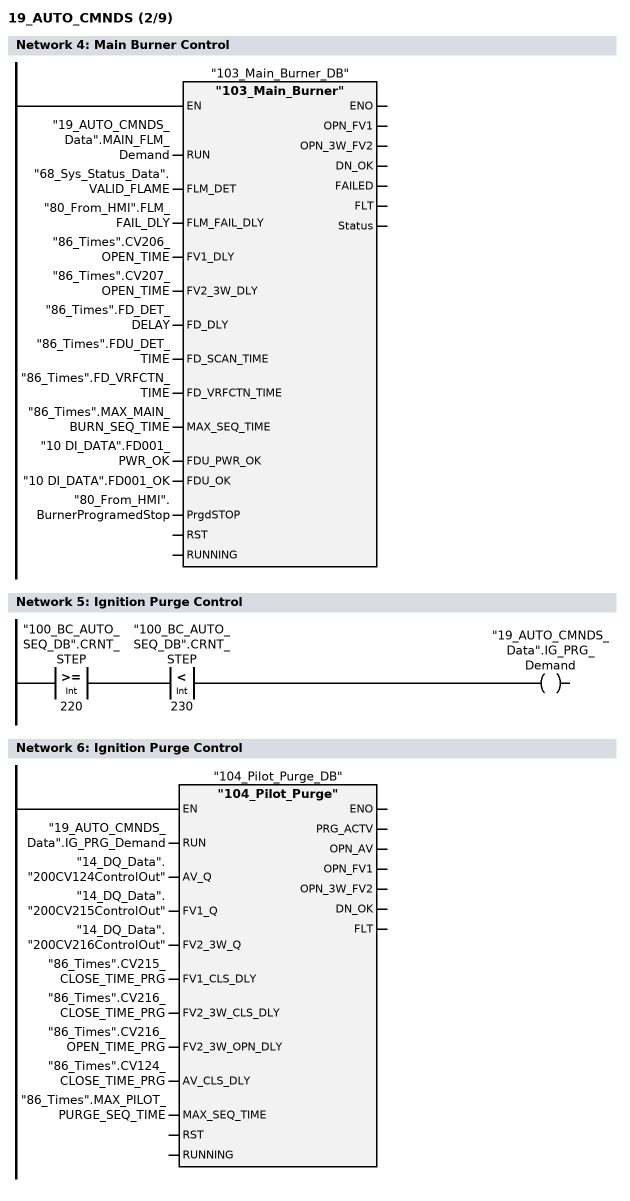
   RUNG wire#powerrail
      "103_Main_Burner_DB"(RUN := "19_AUTO_CMNDS_Data".MAIN_FLM_Demand, FLM_DET := "68_Sys_Status_Data".VALID_FLAME, FLM_FAIL_DLY := "80_From_HMI".FLM_FAIL_DLY, FV1_DLY := "86_Times".CV206_OPEN_TIME, FV2_3W_DLY := "86_Times".CV207_OPEN_TIME, FD_DLY := "86_Times".FD_DET_DELAY, FD_SCAN_TIME := "86_Times".FDU_DET_TIME, FD_VRFCTN_TIME := "86_Times".FD_VRFCTN_TIME, MAX_SEQ_TIME := "86_Times".MAX_MAIN_BURN_SEQ_TIME, FDU_PWR_OK := "10 DI_DATA".FD001_PWR_OK, FDU_OK := "10 DI_DATA".FD001_OK, PrgdSTOP := "80_From_HMI".BurnerProgramedStop, RST :=, RUNNING :=, OPN_FV1 =>, OPN_3W_FV2 =>, DN_OK =>, FAILED =>, FLT =>, Status =>)
   END_RUNG
   // the same network as SCL:
   "103_Main_Burner_DB"(RUN := "19_AUTO_CMNDS_Data".MAIN_FLM_Demand,   // "103_Main_Burner"
                        FLM_DET := "68_Sys_Status_Data".VALID_FLAME,
                        FLM_FAIL_DLY := "80_From_HMI".FLM_FAIL_DLY,
                        FV1_DLY := "86_Times".CV206_OPEN_TIME,
                        FV2_3W_DLY := "86_Times".CV207_OPEN_TIME,
                        FD_DLY := "86_Times".FD_DET_DELAY,
                        FD_SCAN_TIME := "86_Times".FDU_DET_TIME,
                        FD_VRFCTN_TIME := "86_Times".FD_VRFCTN_TIME,
                        MAX_SEQ_TIME := "86_Times".MAX_MAIN_BURN_SEQ_TIME,
                        FDU_PWR_OK := "10 DI_DATA".FD001_PWR_OK,
                        FDU_OK := "10 DI_DATA".FD001_OK,
                        PrgdSTOP := "80_From_HMI".BurnerProgramedStop);
END_REGION

REGION Network 5: Ignition Purge Control
   RUNG wire#powerrail
      { S7_Templates := "SrcType := Int" } GE_Contact(in1 := "100_BC_AUTO_SEQ_DB".CRNT_STEP, in2 := 220)
      { S7_Templates := "SrcType := Int" } LT_Contact(in1 := "100_BC_AUTO_SEQ_DB".CRNT_STEP, in2 := 230)
      Coil( "19_AUTO_CMNDS_Data".IG_PRG_Demand )
   END_RUNG
   // the same network as SCL:
   "19_AUTO_CMNDS_Data".IG_PRG_Demand := ("100_BC_AUTO_SEQ_DB".CRNT_STEP >= 220) AND ("100_BC_AUTO_SEQ_DB".CRNT_STEP < 230);
END_REGION

REGION Network 6: Ignition Purge Control
   RUNG wire#powerrail
      "104_Pilot_Purge_DB"(RUN := "19_AUTO_CMNDS_Data".IG_PRG_Demand, AV_Q := "14_DQ_Data"."200CV124ControlOut", FV1_Q := "14_DQ_Data"."200CV215ControlOut", FV2_3W_Q := "14_DQ_Data"."200CV216ControlOut", FV1_CLS_DLY := "86_Times".CV215_CLOSE_TIME_PRG, FV2_3W_CLS_DLY := "86_Times".CV216_CLOSE_TIME_PRG, FV2_3W_OPN_DLY := "86_Times".CV216_OPEN_TIME_PRG, AV_CLS_DLY := "86_Times".CV124_CLOSE_TIME_PRG, MAX_SEQ_TIME := "86_Times".MAX_PILOT_PURGE_SEQ_TIME, RST :=, RUNNING :=, PRG_ACTV =>, OPN_AV =>, OPN_FV1 =>, OPN_3W_FV2 =>, DN_OK =>, FLT =>)
   END_RUNG
   // the same network as SCL:
   "104_Pilot_Purge_DB"(RUN := "19_AUTO_CMNDS_Data".IG_PRG_Demand,   // "104_Pilot_Purge"
                        AV_Q := "14_DQ_Data"."200CV124ControlOut",
                        FV1_Q := "14_DQ_Data"."200CV215ControlOut",
                        FV2_3W_Q := "14_DQ_Data"."200CV216ControlOut",
                        FV1_CLS_DLY := "86_Times".CV215_CLOSE_TIME_PRG,
                        FV2_3W_CLS_DLY := "86_Times".CV216_CLOSE_TIME_PRG,
                        FV2_3W_OPN_DLY := "86_Times".CV216_OPEN_TIME_PRG,
                        AV_CLS_DLY := "86_Times".CV124_CLOSE_TIME_PRG,
                        MAX_SEQ_TIME := "86_Times".MAX_PILOT_PURGE_SEQ_TIME);
END_REGION

REGION Network 7: Q0.0 - Test pressure valve control CV127
   // True = Open, False = Closed
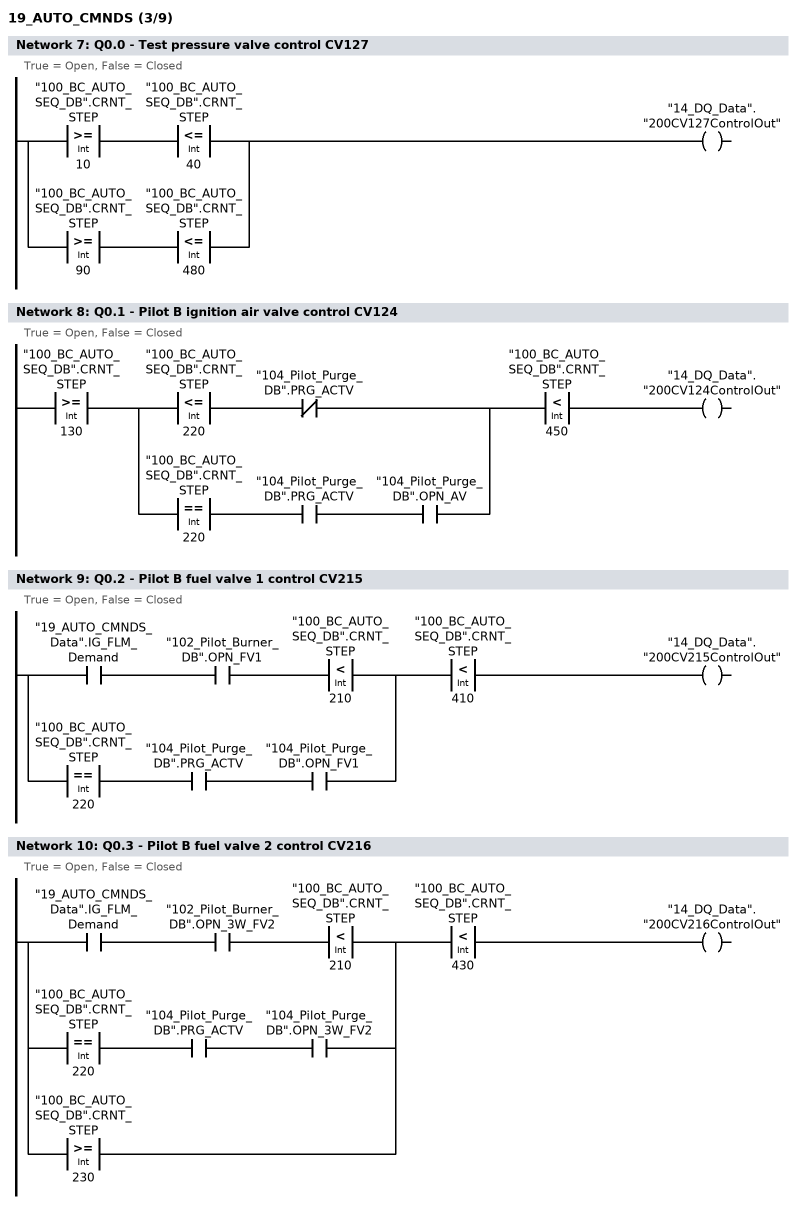
   RUNG wire#powerrail
      { S7_Templates := "SrcType := Int" } GE_Contact(in1 := "100_BC_AUTO_SEQ_DB".CRNT_STEP, in2 := 10)
      { S7_Templates := "SrcType := Int" } LE_Contact(in1 := "100_BC_AUTO_SEQ_DB".CRNT_STEP, in2 := 40)
      wire#w1
      Coil( "14_DQ_Data"."200CV127ControlOut" )
   END_RUNG
   RUNG wire#powerrail
      { S7_Templates := "SrcType := Int" } GE_Contact(in1 := "100_BC_AUTO_SEQ_DB".CRNT_STEP, in2 := 90)
      { S7_Templates := "SrcType := Int" } LE_Contact(in1 := "100_BC_AUTO_SEQ_DB".CRNT_STEP, in2 := 480)
   END_RUNG wire#w1
   // the same network as SCL:
   "14_DQ_Data"."200CV127ControlOut" := (("100_BC_AUTO_SEQ_DB".CRNT_STEP >= 10) AND ("100_BC_AUTO_SEQ_DB".CRNT_STEP <= 40)) OR (("100_BC_AUTO_SEQ_DB".CRNT_STEP >= 90) AND ("100_BC_AUTO_SEQ_DB".CRNT_STEP <= 480));
END_REGION

REGION Network 8: Q0.1 - Pilot B ignition air valve control CV124
   // True = Open, False = Closed
   RUNG wire#powerrail
      { S7_Templates := "SrcType := Int" } GE_Contact(in1 := "100_BC_AUTO_SEQ_DB".CRNT_STEP, in2 := 130)
      wire#w1
      { S7_Templates := "SrcType := Int" } LE_Contact(in1 := "100_BC_AUTO_SEQ_DB".CRNT_STEP, in2 := 220)
      I_Contact( "104_Pilot_Purge_DB".PRG_ACTV )
      wire#w2
      { S7_Templates := "SrcType := Int" } LT_Contact(in1 := "100_BC_AUTO_SEQ_DB".CRNT_STEP, in2 := 450)
      Coil( "14_DQ_Data"."200CV124ControlOut" )
   END_RUNG
   RUNG wire#w1
      { S7_Templates := "SrcType := Int" } EQ_Contact(in1 := "100_BC_AUTO_SEQ_DB".CRNT_STEP, in2 := 220)
      Contact( "104_Pilot_Purge_DB".PRG_ACTV )
      Contact( "104_Pilot_Purge_DB".OPN_AV )
   END_RUNG wire#w2
   // the same network as SCL:
   "14_DQ_Data"."200CV124ControlOut" := ("100_BC_AUTO_SEQ_DB".CRNT_STEP >= 130) AND ((("100_BC_AUTO_SEQ_DB".CRNT_STEP <= 220) AND NOT "104_Pilot_Purge_DB".PRG_ACTV) OR (("100_BC_AUTO_SEQ_DB".CRNT_STEP = 220) AND "104_Pilot_Purge_DB".PRG_ACTV AND "104_Pilot_Purge_DB".OPN_AV)) AND ("100_BC_AUTO_SEQ_DB".CRNT_STEP < 450);
END_REGION

REGION Network 9: Q0.2 - Pilot B fuel valve 1 control CV215
   // True = Open, False = Closed
   RUNG wire#powerrail
      Contact( "19_AUTO_CMNDS_Data".IG_FLM_Demand )
      Contact( "102_Pilot_Burner_DB".OPN_FV1 )
      { S7_Templates := "SrcType := Int" } LT_Contact(in1 := "100_BC_AUTO_SEQ_DB".CRNT_STEP, in2 := 210)
      wire#w1
      { S7_Templates := "SrcType := Int" } LT_Contact(in1 := "100_BC_AUTO_SEQ_DB".CRNT_STEP, in2 := 410)
      Coil( "14_DQ_Data"."200CV215ControlOut" )
   END_RUNG
   RUNG wire#powerrail
      { S7_Templates := "SrcType := Int" } EQ_Contact(in1 := "100_BC_AUTO_SEQ_DB".CRNT_STEP, in2 := 220)
      Contact( "104_Pilot_Purge_DB".PRG_ACTV )
      Contact( "104_Pilot_Purge_DB".OPN_FV1 )
   END_RUNG wire#w1
   // the same network as SCL:
   "14_DQ_Data"."200CV215ControlOut" := (("19_AUTO_CMNDS_Data".IG_FLM_Demand AND "102_Pilot_Burner_DB".OPN_FV1 AND ("100_BC_AUTO_SEQ_DB".CRNT_STEP < 210)) OR (("100_BC_AUTO_SEQ_DB".CRNT_STEP = 220) AND "104_Pilot_Purge_DB".PRG_ACTV AND "104_Pilot_Purge_DB".OPN_FV1)) AND ("100_BC_AUTO_SEQ_DB".CRNT_STEP < 410);
END_REGION

REGION Network 10: Q0.3 - Pilot B fuel valve 2 control CV216
   // True = Open, False = Closed
   RUNG wire#powerrail
      Contact( "19_AUTO_CMNDS_Data".IG_FLM_Demand )
      Contact( "102_Pilot_Burner_DB".OPN_3W_FV2 )
      { S7_Templates := "SrcType := Int" } LT_Contact(in1 := "100_BC_AUTO_SEQ_DB".CRNT_STEP, in2 := 210)
      wire#w1
      { S7_Templates := "SrcType := Int" } LT_Contact(in1 := "100_BC_AUTO_SEQ_DB".CRNT_STEP, in2 := 430)
      Coil( "14_DQ_Data"."200CV216ControlOut" )
   END_RUNG
   RUNG wire#powerrail
      { S7_Templates := "SrcType := Int" } EQ_Contact(in1 := "100_BC_AUTO_SEQ_DB".CRNT_STEP, in2 := 220)
      Contact( "104_Pilot_Purge_DB".PRG_ACTV )
      Contact( "104_Pilot_Purge_DB".OPN_3W_FV2 )
   END_RUNG wire#w1
   RUNG wire#powerrail
      { S7_Templates := "SrcType := Int" } GE_Contact(in1 := "100_BC_AUTO_SEQ_DB".CRNT_STEP, in2 := 230)
   END_RUNG wire#w1
   // the same network as SCL:
   "14_DQ_Data"."200CV216ControlOut" := (("19_AUTO_CMNDS_Data".IG_FLM_Demand AND "102_Pilot_Burner_DB".OPN_3W_FV2 AND ("100_BC_AUTO_SEQ_DB".CRNT_STEP < 210)) OR (("100_BC_AUTO_SEQ_DB".CRNT_STEP = 220) AND "104_Pilot_Purge_DB".PRG_ACTV AND "104_Pilot_Purge_DB".OPN_3W_FV2) OR ("100_BC_AUTO_SEQ_DB".CRNT_STEP >= 230)) AND ("100_BC_AUTO_SEQ_DB".CRNT_STEP < 430);
END_REGION

REGION Network 11: Q0.4 - Main B atom air valve control CV114
   // True = Open, False = Closed
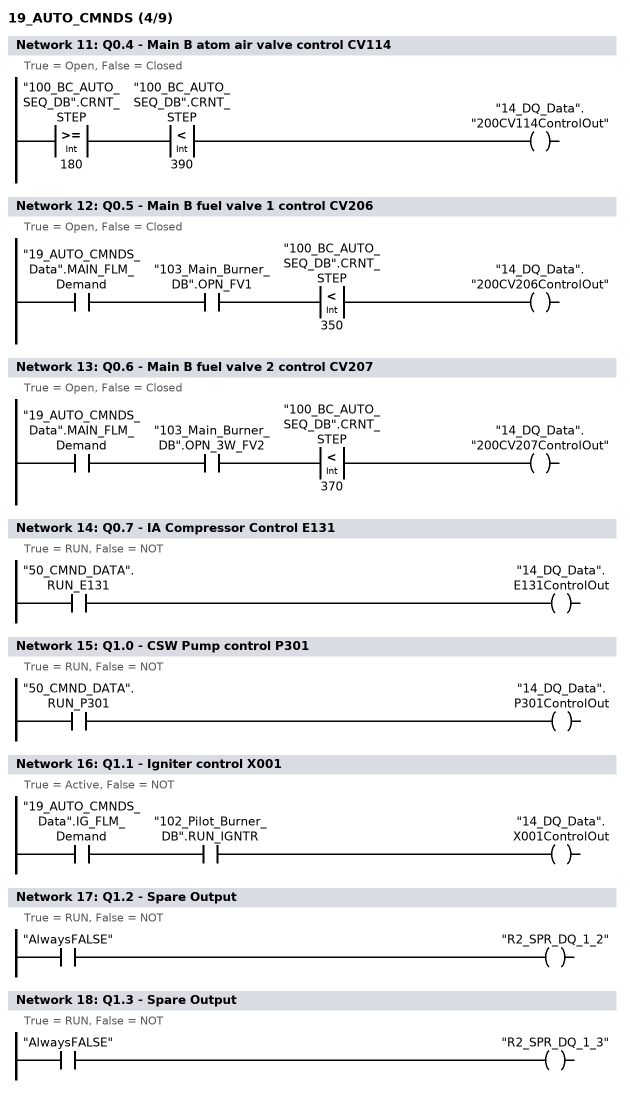
   RUNG wire#powerrail
      { S7_Templates := "SrcType := Int" } GE_Contact(in1 := "100_BC_AUTO_SEQ_DB".CRNT_STEP, in2 := 180)
      { S7_Templates := "SrcType := Int" } LT_Contact(in1 := "100_BC_AUTO_SEQ_DB".CRNT_STEP, in2 := 390)
      Coil( "14_DQ_Data"."200CV114ControlOut" )
   END_RUNG
   // the same network as SCL:
   "14_DQ_Data"."200CV114ControlOut" := ("100_BC_AUTO_SEQ_DB".CRNT_STEP >= 180) AND ("100_BC_AUTO_SEQ_DB".CRNT_STEP < 390);
END_REGION

REGION Network 12: Q0.5 - Main B fuel valve 1 control CV206
   // True = Open, False = Closed
   RUNG wire#powerrail
      Contact( "19_AUTO_CMNDS_Data".MAIN_FLM_Demand )
      Contact( "103_Main_Burner_DB".OPN_FV1 )
      { S7_Templates := "SrcType := Int" } LT_Contact(in1 := "100_BC_AUTO_SEQ_DB".CRNT_STEP, in2 := 350)
      Coil( "14_DQ_Data"."200CV206ControlOut" )
   END_RUNG
   // the same network as SCL:
   "14_DQ_Data"."200CV206ControlOut" := "19_AUTO_CMNDS_Data".MAIN_FLM_Demand AND "103_Main_Burner_DB".OPN_FV1 AND ("100_BC_AUTO_SEQ_DB".CRNT_STEP < 350);
END_REGION

REGION Network 13: Q0.6 - Main B fuel valve 2 control CV207
   // True = Open, False = Closed
   RUNG wire#powerrail
      Contact( "19_AUTO_CMNDS_Data".MAIN_FLM_Demand )
      Contact( "103_Main_Burner_DB".OPN_3W_FV2 )
      { S7_Templates := "SrcType := Int" } LT_Contact(in1 := "100_BC_AUTO_SEQ_DB".CRNT_STEP, in2 := 370)
      Coil( "14_DQ_Data"."200CV207ControlOut" )
   END_RUNG
   // the same network as SCL:
   "14_DQ_Data"."200CV207ControlOut" := "19_AUTO_CMNDS_Data".MAIN_FLM_Demand AND "103_Main_Burner_DB".OPN_3W_FV2 AND ("100_BC_AUTO_SEQ_DB".CRNT_STEP < 370);
END_REGION

REGION Network 14: Q0.7 - IA Compressor Control E131
   // True = RUN, False = NOT
   RUNG wire#powerrail
      Contact( "50_CMND_DATA".RUN_E131 )
      Coil( "14_DQ_Data".E131ControlOut )
   END_RUNG
   // the same network as SCL:
   "14_DQ_Data".E131ControlOut := "50_CMND_DATA".RUN_E131;
END_REGION

REGION Network 15: Q1.0 - CSW Pump control P301
   // True = RUN, False = NOT
   RUNG wire#powerrail
      Contact( "50_CMND_DATA".RUN_P301 )
      Coil( "14_DQ_Data".P301ControlOut )
   END_RUNG
   // the same network as SCL:
   "14_DQ_Data".P301ControlOut := "50_CMND_DATA".RUN_P301;
END_REGION

REGION Network 16: Q1.1 - Igniter control X001
   // True = Active, False = NOT
   RUNG wire#powerrail
      Contact( "19_AUTO_CMNDS_Data".IG_FLM_Demand )
      Contact( "102_Pilot_Burner_DB".RUN_IGNTR )
      Coil( "14_DQ_Data".X001ControlOut )
   END_RUNG
   // the same network as SCL:
   "14_DQ_Data".X001ControlOut := "19_AUTO_CMNDS_Data".IG_FLM_Demand AND "102_Pilot_Burner_DB".RUN_IGNTR;
END_REGION

REGION Network 17: Q1.2 - Spare Output
   // True = RUN, False = NOT
   RUNG wire#powerrail
      Contact( "AlwaysFALSE" )
      Coil( "R2_SPR_DQ_1_2" )
   END_RUNG
   // the same network as SCL:
   "R2_SPR_DQ_1_2" := "AlwaysFALSE";
END_REGION

REGION Network 18: Q1.3 - Spare Output
   // True = RUN, False = NOT
   RUNG wire#powerrail
      Contact( "AlwaysFALSE" )
      Coil( "R2_SPR_DQ_1_3" )
   END_RUNG
   // the same network as SCL:
   "R2_SPR_DQ_1_3" := "AlwaysFALSE";
END_REGION

REGION Network 19: Q1.4 - Spare Output
   // True = RUN, False = NOT
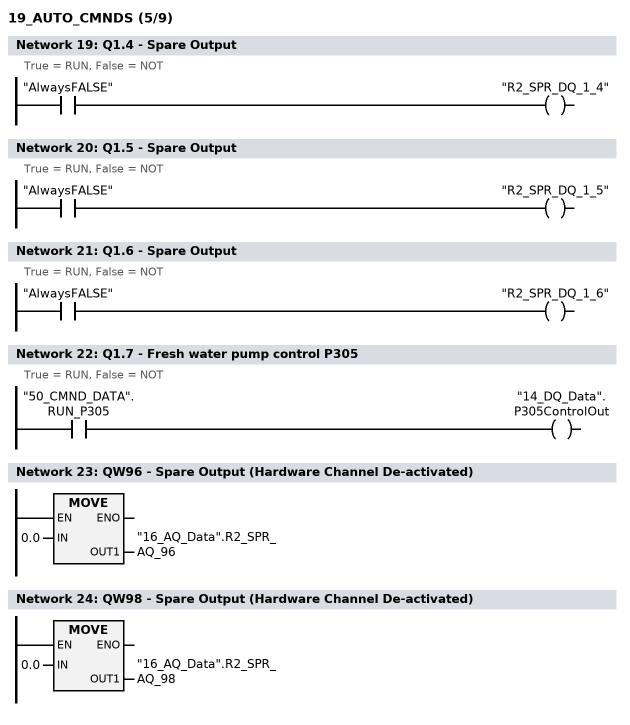
   RUNG wire#powerrail
      Contact( "AlwaysFALSE" )
      Coil( "R2_SPR_DQ_1_4" )
   END_RUNG
   // the same network as SCL:
   "R2_SPR_DQ_1_4" := "AlwaysFALSE";
END_REGION

REGION Network 20: Q1.5 - Spare Output
   // True = RUN, False = NOT
   RUNG wire#powerrail
      Contact( "AlwaysFALSE" )
      Coil( "R2_SPR_DQ_1_5" )
   END_RUNG
   // the same network as SCL:
   "R2_SPR_DQ_1_5" := "AlwaysFALSE";
END_REGION

REGION Network 21: Q1.6 - Spare Output
   // True = RUN, False = NOT
   RUNG wire#powerrail
      Contact( "AlwaysFALSE" )
      Coil( "R2_SPR_DQ_1_6" )
   END_RUNG
   // the same network as SCL:
   "R2_SPR_DQ_1_6" := "AlwaysFALSE";
END_REGION

REGION Network 22: Q1.7 - Fresh water pump control P305
   // True = RUN, False = NOT
   RUNG wire#powerrail
      Contact( "50_CMND_DATA".RUN_P305 )
      Coil( "14_DQ_Data".P305ControlOut )
   END_RUNG
   // the same network as SCL:
   "14_DQ_Data".P305ControlOut := "50_CMND_DATA".RUN_P305;
END_REGION

REGION Network 23: QW96 - Spare Output (Hardware Channel De-activated)
   RUNG wire#powerrail
      Move(in := 0.0, out1 => "16_AQ_Data".R2_SPR_AQ_96)
   END_RUNG
   // the same network as SCL:
   "16_AQ_Data".R2_SPR_AQ_96 := 0.0;
END_REGION

REGION Network 24: QW98 - Spare Output (Hardware Channel De-activated)
   RUNG wire#powerrail
      Move(in := 0.0, out1 => "16_AQ_Data".R2_SPR_AQ_98)
   END_RUNG
   // the same network as SCL:
   "16_AQ_Data".R2_SPR_AQ_98 := 0.0;
END_REGION

REGION Network 25: QW100 - Main Fuel Reg Valve Control CV203 (For Main Burn Start)
   // Changed from 20 to 230 at 160 to230 for test
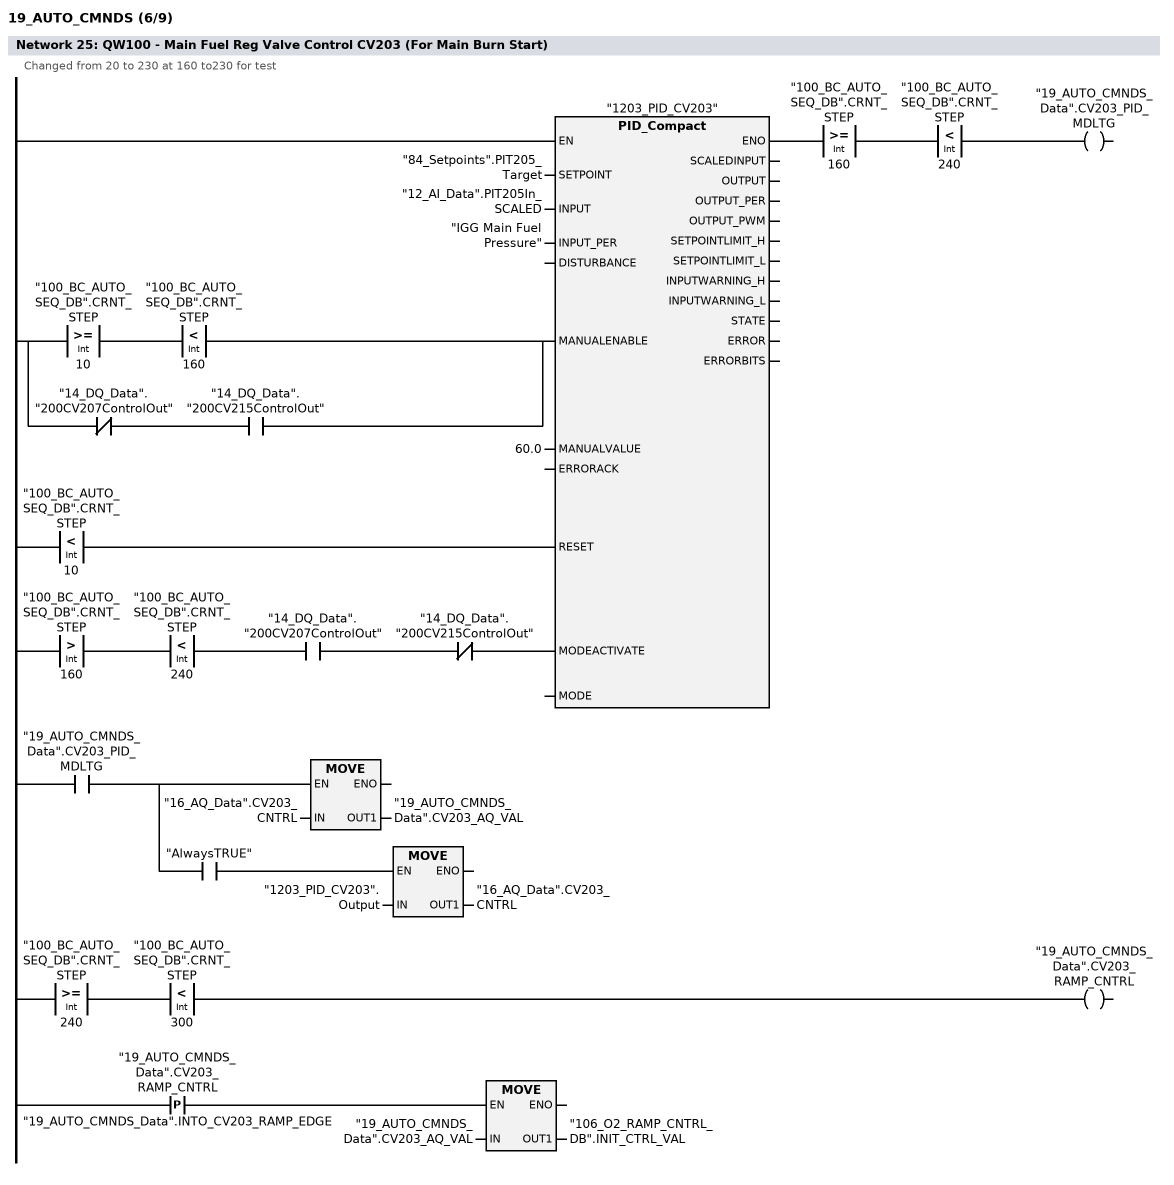
   // ENO of a box is taken as its EN; it also drops when the box reports an error
   "1203_PID_CV203"(Setpoint := "84_Setpoints".PIT205_Target,   // PID_Compact
                    Input := "12_AI_Data".PIT205In_SCALED,
                    Input_PER := "IGG Main Fuel Pressure",
                    ManualEnable := (("100_BC_AUTO_SEQ_DB".CRNT_STEP >= 10) AND ("100_BC_AUTO_SEQ_DB".CRNT_STEP < 160)) OR (NOT "14_DQ_Data"."200CV207ControlOut" AND "14_DQ_Data"."200CV215ControlOut"),
                    ManualValue := 60.0,
                    Reset := "100_BC_AUTO_SEQ_DB".CRNT_STEP < 10,
                    ModeActivate := ("100_BC_AUTO_SEQ_DB".CRNT_STEP > 160) AND ("100_BC_AUTO_SEQ_DB".CRNT_STEP < 240) AND "14_DQ_Data"."200CV207ControlOut" AND NOT "14_DQ_Data"."200CV215ControlOut");
   "19_AUTO_CMNDS_Data".CV203_PID_MDLTG := ("100_BC_AUTO_SEQ_DB".CRNT_STEP >= 160) AND ("100_BC_AUTO_SEQ_DB".CRNT_STEP < 240);
   IF "19_AUTO_CMNDS_Data".CV203_PID_MDLTG THEN
       "19_AUTO_CMNDS_Data".CV203_AQ_VAL := "16_AQ_Data".CV203_CNTRL;
   END_IF;
   IF "19_AUTO_CMNDS_Data".CV203_PID_MDLTG AND "AlwaysTRUE" THEN
       "16_AQ_Data".CV203_CNTRL := "1203_PID_CV203".Output;
   END_IF;
   "19_AUTO_CMNDS_Data".CV203_RAMP_CNTRL := ("100_BC_AUTO_SEQ_DB".CRNT_STEP >= 240) AND ("100_BC_AUTO_SEQ_DB".CRNT_STEP < 300);
   #_w1 := "19_AUTO_CMNDS_Data".CV203_RAMP_CNTRL AND NOT "19_AUTO_CMNDS_Data".INTO_CV203_RAMP_EDGE;   // rising edge of "19_AUTO_CMNDS_Data".CV203_RAMP_CNTRL
   "19_AUTO_CMNDS_Data".INTO_CV203_RAMP_EDGE := "19_AUTO_CMNDS_Data".CV203_RAMP_CNTRL;
   IF #_w1 THEN "106_O2_RAMP_CNTRL_DB".INIT_CTRL_VAL := "19_AUTO_CMNDS_Data".CV203_AQ_VAL; END_IF;
END_REGION

REGION Network 26: QW100 - Main Fuel Reg Valve Control CV203 (Ramp for O2)
   // To delete this FB106 when time for testing available
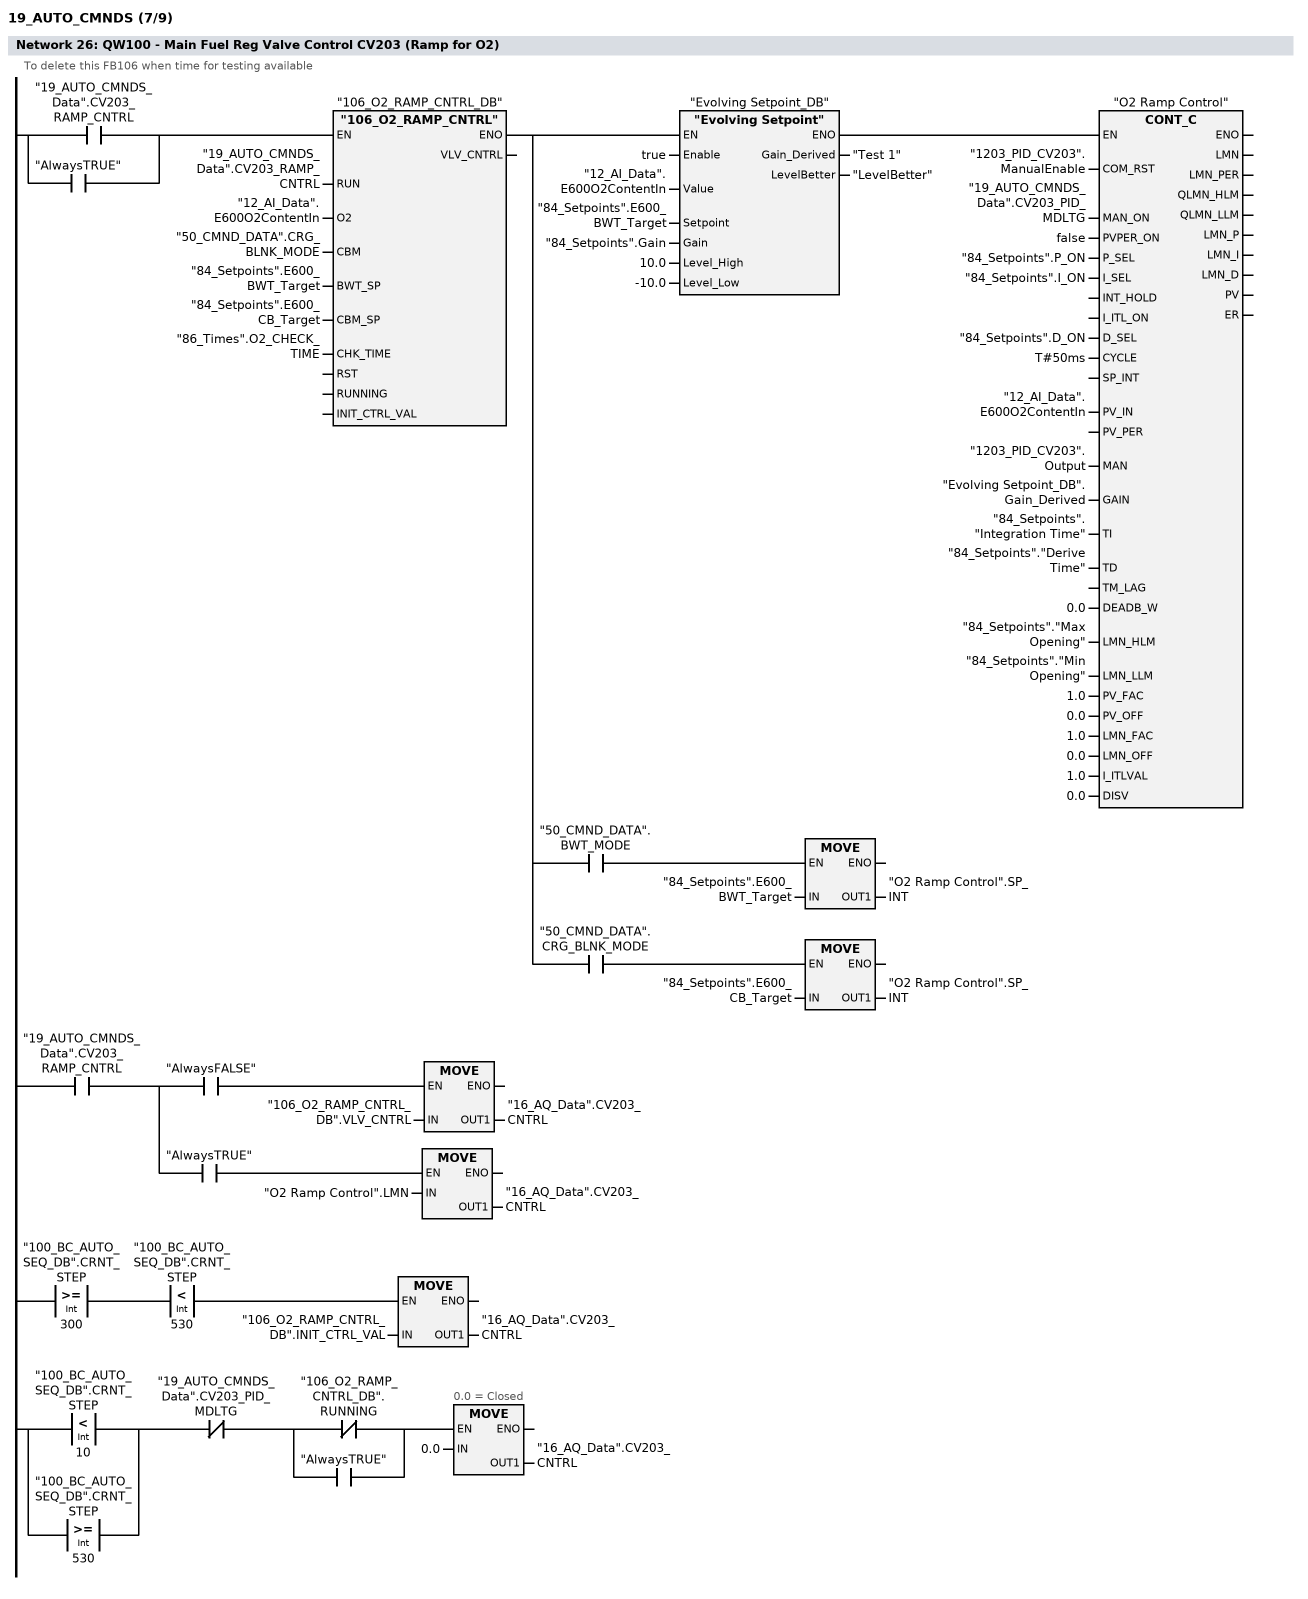
   "106_O2_RAMP_CNTRL_DB"(EN := "19_AUTO_CMNDS_Data".CV203_RAMP_CNTRL OR "AlwaysTRUE",   // "106_O2_RAMP_CNTRL"
                          RUN := "19_AUTO_CMNDS_Data".CV203_RAMP_CNTRL,
                          O2 := "12_AI_Data".E600O2ContentIn,
                          CBM := "50_CMND_DATA".CRG_BLNK_MODE,
                          BWT_SP := "84_Setpoints".E600_BWT_Target,
                          CBM_SP := "84_Setpoints".E600_CB_Target,
                          CHK_TIME := "86_Times".O2_CHECK_TIME,
                          ENO => #_w1);
   "Evolving Setpoint_DB"(EN := #_w1,   // "Evolving Setpoint"
                          Enable := true,
                          Value := "12_AI_Data".E600O2ContentIn,
                          Setpoint := "84_Setpoints".E600_BWT_Target,
                          Gain := "84_Setpoints".Gain,
                          Level_High := 10.0,
                          Level_Low := -10.0,
                          Gain_Derived => "Test 1",
                          LevelBetter => "LevelBetter",
                          ENO => #_w2);
   IF #_w2 THEN
       "O2 Ramp Control"(COM_RST := "1203_PID_CV203".ManualEnable,   // CONT_C
                         MAN_ON := "19_AUTO_CMNDS_Data".CV203_PID_MDLTG,
                         PVPER_ON := false,
                         P_SEL := "84_Setpoints".P_ON,
                         I_SEL := "84_Setpoints".I_ON,
                         D_SEL := "84_Setpoints".D_ON,
                         CYCLE := T#50ms,
                         PV_IN := "12_AI_Data".E600O2ContentIn,
                         MAN := "1203_PID_CV203".Output,
                         GAIN := "Evolving Setpoint_DB".Gain_Derived,
                         TI := "84_Setpoints"."Integration Time",
                         TD := "84_Setpoints"."Derive Time",
                         DEADB_W := 0.0,
                         LMN_HLM := "84_Setpoints"."Max Opening",
                         LMN_LLM := "84_Setpoints"."Min Opening",
                         PV_FAC := 1.0,
                         PV_OFF := 0.0,
                         LMN_FAC := 1.0,
                         LMN_OFF := 0.0,
                         I_ITLVAL := 1.0,
                         DISV := 0.0);
   END_IF;
   IF #_w1 AND "50_CMND_DATA".BWT_MODE THEN
       "O2 Ramp Control".SP_INT := "84_Setpoints".E600_BWT_Target;
   END_IF;
   IF #_w1 AND "50_CMND_DATA".CRG_BLNK_MODE THEN
       "O2 Ramp Control".SP_INT := "84_Setpoints".E600_CB_Target;
   END_IF;
   IF "19_AUTO_CMNDS_Data".CV203_RAMP_CNTRL AND "AlwaysFALSE" THEN
       "16_AQ_Data".CV203_CNTRL := "106_O2_RAMP_CNTRL_DB".VLV_CNTRL;
   END_IF;
   IF "19_AUTO_CMNDS_Data".CV203_RAMP_CNTRL AND "AlwaysTRUE" THEN
       "16_AQ_Data".CV203_CNTRL := "O2 Ramp Control".LMN;
   END_IF;
   IF ("100_BC_AUTO_SEQ_DB".CRNT_STEP >= 300) AND ("100_BC_AUTO_SEQ_DB".CRNT_STEP < 530) THEN
       "16_AQ_Data".CV203_CNTRL := "106_O2_RAMP_CNTRL_DB".INIT_CTRL_VAL;
   END_IF;
   IF (("100_BC_AUTO_SEQ_DB".CRNT_STEP < 10) OR ("100_BC_AUTO_SEQ_DB".CRNT_STEP >= 530)) AND NOT "19_AUTO_CMNDS_Data".CV203_PID_MDLTG AND (NOT "106_O2_RAMP_CNTRL_DB".RUNNING OR "AlwaysTRUE") THEN
       "16_AQ_Data".CV203_CNTRL := 0.0;   // 0.0 = Closed
   END_IF;
END_REGION

REGION Network 27: CV111 setpoints
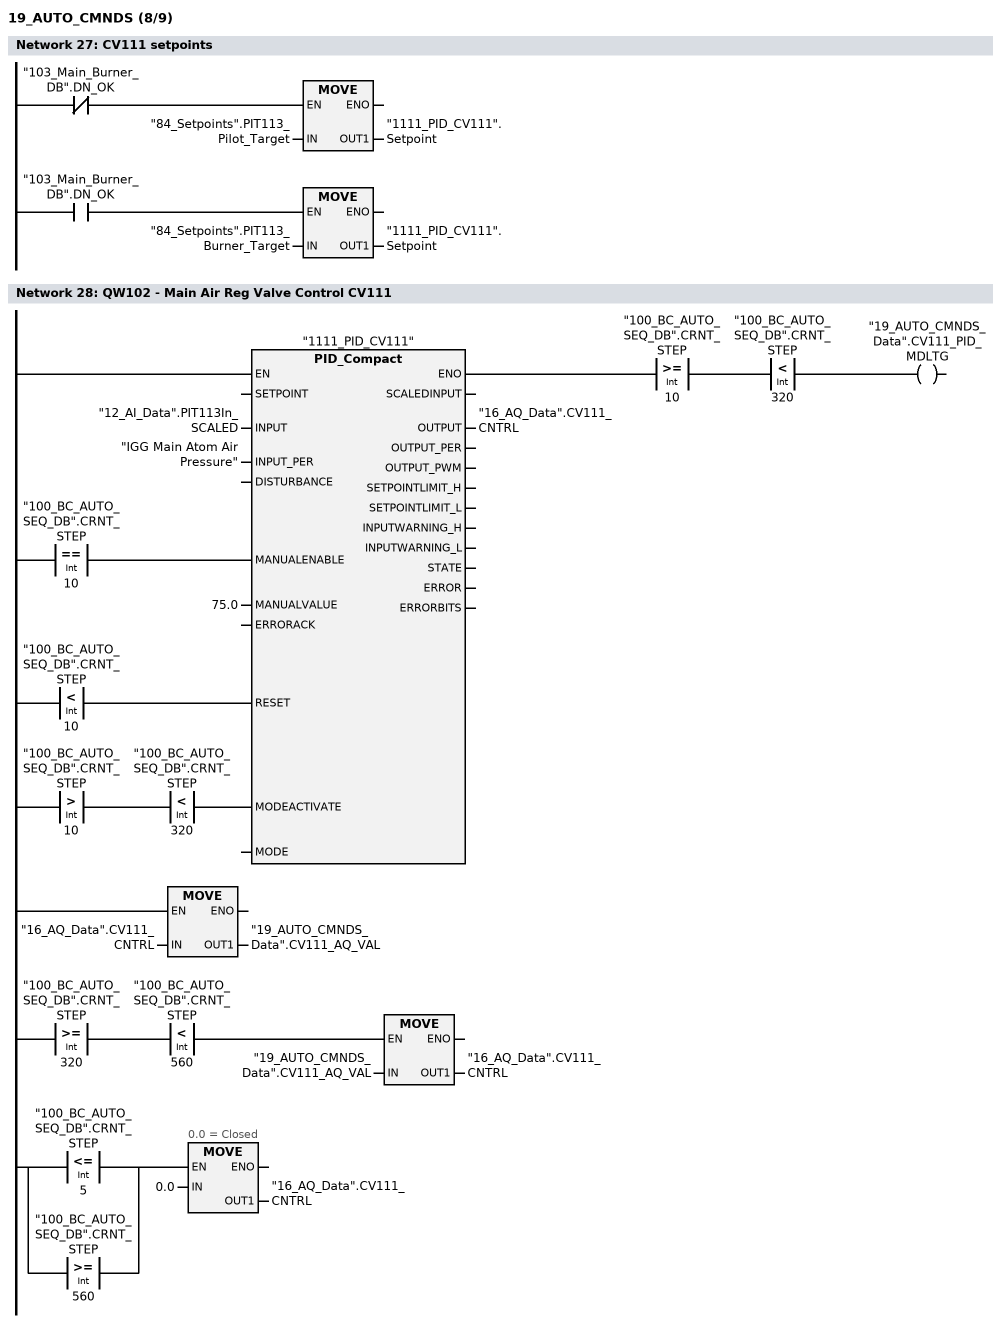
   RUNG wire#powerrail
      I_Contact( "103_Main_Burner_DB".DN_OK )
      Move(in := "84_Setpoints".PIT113_Pilot_Target, out1 => "1111_PID_CV111".Setpoint)
   END_RUNG
   RUNG wire#powerrail
      Contact( "103_Main_Burner_DB".DN_OK )
      Move(in := "84_Setpoints".PIT113_Burner_Target, out1 => "1111_PID_CV111".Setpoint)
   END_RUNG
   // the same network as SCL:
   IF NOT "103_Main_Burner_DB".DN_OK THEN
       "1111_PID_CV111".Setpoint := "84_Setpoints".PIT113_Pilot_Target;
   END_IF;
   IF "103_Main_Burner_DB".DN_OK THEN
       "1111_PID_CV111".Setpoint := "84_Setpoints".PIT113_Burner_Target;
   END_IF;
END_REGION

REGION Network 28: QW102 - Main Air Reg Valve Control CV111
   // ENO of a box is taken as its EN; it also drops when the box reports an error
   "1111_PID_CV111"(Input := "12_AI_Data".PIT113In_SCALED,   // PID_Compact
                    Input_PER := "IGG Main Atom Air Pressure",
                    ManualEnable := "100_BC_AUTO_SEQ_DB".CRNT_STEP = 10,
                    ManualValue := 75.0,
                    Reset := "100_BC_AUTO_SEQ_DB".CRNT_STEP < 10,
                    ModeActivate := ("100_BC_AUTO_SEQ_DB".CRNT_STEP > 10) AND ("100_BC_AUTO_SEQ_DB".CRNT_STEP < 320),
                    Output => "16_AQ_Data".CV111_CNTRL);
   "19_AUTO_CMNDS_Data".CV111_PID_MDLTG := ("100_BC_AUTO_SEQ_DB".CRNT_STEP >= 10) AND ("100_BC_AUTO_SEQ_DB".CRNT_STEP < 320);
   "19_AUTO_CMNDS_Data".CV111_AQ_VAL := "16_AQ_Data".CV111_CNTRL;
   IF ("100_BC_AUTO_SEQ_DB".CRNT_STEP >= 320) AND ("100_BC_AUTO_SEQ_DB".CRNT_STEP < 560) THEN
       "16_AQ_Data".CV111_CNTRL := "19_AUTO_CMNDS_Data".CV111_AQ_VAL;
   END_IF;
   IF ("100_BC_AUTO_SEQ_DB".CRNT_STEP <= 5) OR ("100_BC_AUTO_SEQ_DB".CRNT_STEP >= 560) THEN
       "16_AQ_Data".CV111_CNTRL := 0.0;   // 0.0 = Closed
   END_IF;
END_REGION

REGION Network 30: IGG - Pilot Burner Confirmed
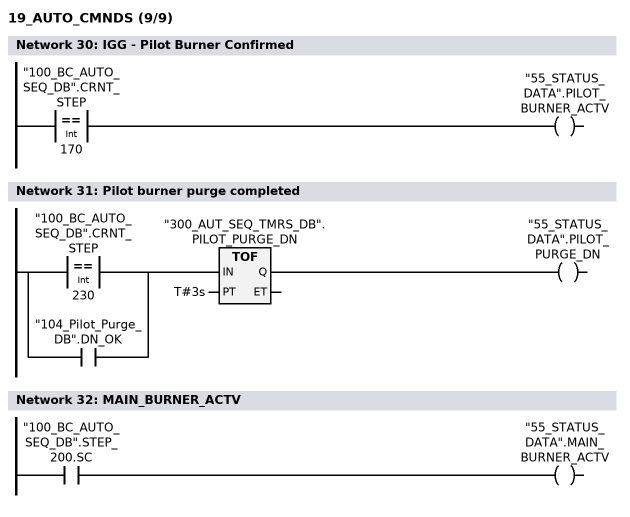
   RUNG wire#powerrail
      { S7_Templates := "SrcType := Int" } EQ_Contact(in1 := "100_BC_AUTO_SEQ_DB".CRNT_STEP, in2 := 170)
      Coil( "55_STATUS_DATA".PILOT_BURNER_ACTV )
   END_RUNG
   // the same network as SCL:
   "55_STATUS_DATA".PILOT_BURNER_ACTV := "100_BC_AUTO_SEQ_DB".CRNT_STEP = 170;
END_REGION

REGION Network 31: Pilot burner purge completed
   "300_AUT_SEQ_TMRS_DB".PILOT_PURGE_DN.TOF(IN := ("100_BC_AUTO_SEQ_DB".CRNT_STEP = 230) OR "104_Pilot_Purge_DB".DN_OK,
                           PT := T#3s);
   "55_STATUS_DATA".PILOT_PURGE_DN := "300_AUT_SEQ_TMRS_DB".PILOT_PURGE_DN.Q;
END_REGION

REGION Network 32: MAIN_BURNER_ACTV
   RUNG wire#powerrail
      Contact( "100_BC_AUTO_SEQ_DB".STEP_200.SC )
      Coil( "55_STATUS_DATA".MAIN_BURNER_ACTV )
   END_RUNG
   // the same network as SCL:
   "55_STATUS_DATA".MAIN_BURNER_ACTV := "100_BC_AUTO_SEQ_DB".STEP_200.SC;
END_REGION
END_FUNCTION

// folder: 100 - 199 Automatic Sequencing

FUNCTION_BLOCK "100_BC_AUTO_SEQ"   // FB100, LAD
TITLE = Automatic Sequence
{ S7_Optimized_Access := 'TRUE' }
AUTHOR : JRS